recipe "配方_5": 总捻度 <- "ST_HMI_Var_HMI_r64NianDu_all", 支数 <- "ST_HMI_Var_HMI_r64ZhiShu_ChengSha", 牵伸捻度匹配值 <- "ST_HMI_Var_HMI_r64NianDu_QianShen_Best", 出车速度 <- "ST_HMI_Var_HMI_r64Velocity_ChuChe", 追捻开始捻度 <- "ST_HMI_Var_HMI_r64NianDu_1", 追捻锭子速度 <- "ST_HMI_Var_HMI_r64NianSu_2", 捻缩开始捻度 <- "ST_HMI_Var_HMI_r64NianDu_NianSuo", 捻缩距离 <- "ST_HMI_Var_HMI_r64Position_NianSuo", 追捻启用开关 <- "ST_HMI_Var_HMI_boNianDu_3"

screen "保养提示" 1280x733, template "模板_2"
   on GenerateScreen: SetTag("变量_100", 6)
   Button "HmiScreenItemData_1" at 1116,65 size 159x60; TextOn '向后 / 後向き / 뒤로'; TextOff '向后 / 後向き / 뒤로'
      on Release: ActivateScreen("自动画面", 0)
   TextField "文本域_6" at 16,8 size 995x720; Text '1.锭子油更换:每隔 天,更换一次 2.龙带传动部分12个黄油嘴，加黄油（耐高温、高速、高负荷） 3.龙带压紧器，加黄油（耐高温 、高速、高负荷） 4.弓轴滚针轴承，每年加一次黄油 5.TC龙带，每两年清洗一次，水温小于15℃，阴凉通风处晾干 6.锭子传动同步带8M-2272 检查维护 7.控制柜清洁，三个月一次,用吸吹风机来吸内部粉尘 8.锭子电机风扇绕毛清理，两个月清理一次 9.其他，走车同步带轮、走车走轮绕毛定期检查清理 1．スピンドル油交換 日,更换一次 2. タンジェントベルト伝動部12ヶ所グリスニップルに、グリス注油（耐高温・高速・高負荷） 3．タンジェントベルトのテークアップ装置にグリス注油（耐高温・高速・高負荷） 4．フォーラーシャフトのニードルベアリングに、年一回グリス注油 5．タンジェンシャルベルトを2年ごとに一回ぬるま湯（水温15℃）で洗い、かげ干しを行う。 6．スピンドル駆動タイミングベルト（８Ｍ－２２７２）点検勧奨 7．コントロールボックスを清潔にし、換気扇の粉塵を三か月ごとに吹き飛ばす。 8．锭子电机风扇绕毛清理，两个月清理一次 9．其他，走车同步带轮、走车走轮绕毛定期检查清理 1. 스핀들오일 교체: 일 간격으로 한번씩 교체한다. 2. tangential belt 전동부분12개 그리스 니플에 그리스 주입(내고온,고속,고부하) 3. 콘택트롤러에그리스 주입한다.(내고온,고속,고부하) 4. 호랑축 니들 베어링은 1년에한번씩 그리스 주입한다. 5. TCtangential belt는2년에 한번씩 청소하고 수온은 15℃이하여야 하며 서늘하고 통 풍이 잘되는곳에 말린다. 6. 스핀들 전동 타이밍벨트8M-2272를점검,유지보수한다. 7. 제어함 청소는 3개월에 한번씩 하고 흡입 송풍기로 내부 분진을 흡입한다. 8. 스핀들 모터팬감긴 원료（绕毛）청소는 2개월에 한번씩한다. 9. 기타 캐리지타이밍풀리,캐리지유동륜은정기적으로 감긴 원료(绕毛)점검,정리한다.'
   IOField "IO 域_3" at 906,98 size 65x39; FormatPattern 999
      ProcessValue <- "ST_Maintenance_g_u16_1_Times_OilChange_DingZi"
   IOField "IO 域_4" at 906,143 size 65x39; FormatPattern 999
      ProcessValue <- "ST_Maintenance_g_u16_2_Times_LongDai_HuangYouZui"
   IOField "IO 域_5" at 906,189 size 65x40; FormatPattern 999
      ProcessValue <- "ST_Maintenance_g_u16_3_Times_LongDai_YaJinQi"
   IOField "IO 域_6" at 906,236 size 65x39; FormatPattern 999
      ProcessValue <- "ST_Maintenance_g_u16_4_Times_GongZhou_Bearing"
   IOField "IO 域_7" at 906,282 size 65x39; FormatPattern 999
      ProcessValue <- "ST_Maintenance_g_u16_5_Times_LongDai_Clean"
   IOField "IO 域_8" at 906,328 size 65x40; FormatPattern 999
      ProcessValue <- "ST_Maintenance_g_u16_6_Times_DingZi_ChuanDong"
   IOField "IO 域_9" at 906,375 size 65x39; FormatPattern 999
      ProcessValue <- "ST_Maintenance_g_u16_7_Times_ControlBox_Clean"
   IOField "IO 域_10" at 906,421 size 65x39; FormatPattern 999
      ProcessValue <- "ST_Maintenance_g_u16_8_Times_DingZi_Fan"
   IOField "IO 域_1" at 258,96 size 66x39; Authorization "User administration"; FormatPattern 999
      ProcessValue <- "ST_Maintenance_g_u16_TimeInterval_OilChange"
   IOField "IO 域_2" at 486,15 size 65x39; Authorization "User administration"; FormatPattern 999
      ProcessValue <- "ST_Maintenance_g_u16_TimeReminder_Maintennance"
   TextField "文本域_4" at 334,19 size 149x32; Text '保养提醒持续 / 保全提醒 / 유지보수 알림'
   TextField "文本域_5" at 563,19 size 48x32; Text '天 / 日 / 일'
   Button "OBJECT_124" at 396,610 size 160x66; TextOn '罗拉关 / 롤러 off'; TextOff '罗拉开关 / EXIT / ローラースイッチ / 롤러 스위치'; Authorization "Operate_5"
      on Release: InvertBit("ST_Main_Var_ST_LuoLaSwitch")
      Appearance <- "ST_Main_Var_ST_LuoLaSwitch"
   TextField "文本域_1" at 40,56 size 149x32; Text '保养项目 / 保全項目 / 유지보수 항목'
   TextField "文本域_2" at 850,56 size 149x32; Text '保养次数 / 保全回数 / 유지보수 횟수'

screen "报警画面" 1280x733, template "模板_2"
   on GenerateScreen: SetTag("变量_100", 5)
   Button "HmiScreenItemData_1" at 1112,90 size 159x60; TextOn '向后 / 後向き / 뒤로'; TextOff '向后 / 後向き / 뒤로'
      on Release: function_efd93a16()
   Button "HmiScreenItemData_2" at 1112,224 size 159x60; TextOn '向后 / 後向き / 뒤로'; TextOff '报警记录 / 警報記録 / 경보알람기록'
      on Release: ActivateScreen("报警记录", 0)
   Button "HmiScreenItemData_3" at 1112,360 size 159x60; TextOn '向后 / 後向き / 뒤로'; TextOff '自动画面 / 自動画面 / 자동화면'
      on Release: ActivateScreen("自动画面", 0)
   AlarmView "报警视图_1" at 3,3 size 1101x728

screen "报警记录" 1280x733, template "模板_2"
   on GenerateScreen: SetTag("变量_100", 16)
   AlarmView "报警视图_1" at 3,2 size 1105x729; ColumnTextDevice 'D425 / PLC / API / ПЛК'
   Button "HmiScreenItemData_2" at 1118,71 size 159x60; TextOn '向后 / 後向き / 뒤로'; TextOff '向后 / 後向き / 뒤로'
      on Release: ActivateScreen("报警画面", 0)

screen "生头画面" 1280x733, template "模板_2"
   on GenerateScreen: SetTag("变量_100", 4)
   Button "HmiScreenItemData_1" at 1118,192 size 159x60; TextOn '向后 / 後向き / 뒤로'; TextOff '向后 / 後向き / 뒤로'
      on Release: ActivateScreen("自动画面", 0)
   Button "OBJECT_107" at 864,104 size 200x65; TextOff '手动 / EXIT / 手動 / 수동'
      on Press: SetTag("ST_Main_Var_g_i16_Mode_Selected", 4)
      Appearance <- "ST_Main_Var_g_bo_Mode_Enabled_Manual"
   Button "OBJECT_108" at 864,192 size 200x65; TextOff '空锭(先插管) EXIT 空鍾（糸管挿入済み） 아이들 스핀들 (먼저 보빈관을 삼입)'
      on Release: ResetBit("ST_HMI_Var_HMI_bo_KongDingShengTou")
      on Press: SetBit("ST_HMI_Var_HMI_bo_KongDingShengTou")
      Appearance <- "ST_HMI_Var_HMI_i16_ShengTou_Select"
   Button "OBJECT_106" at 1041,4 size 238x39; TextOff '手动 / EXIT / 手動 / 수동'; TextList "mode_enabled_1"
      ProcessValue <- "ST_Main_Var_g_i16_Mode_Enabled"
      Appearance <- "ST_Main_Var_g_i16_Mode_Enabled"
   TextField "Text Field_45" at 370,139 size 151x47; Text '实际牵伸: / 実際ドラフト: / 실제 드라프트:'
   TextField "Text Field_46" at 370,205 size 151x47; Text '分散牵伸: / 分散ドラフト: / 스핀들 드라프트:'
   TextField "Text Field_47" at 370,270 size 151x47; Text '走车位置: / キャレージ位置: / 캐리지위치:'
   Button "OBJECT_111" at 1041,43 size 238x40; TextOff '手动 / EXIT / 手動 / 수동'; TextList "KongDing_status#mig1"
      Visibility <- "ST_Main_Var_g_bo_Mode_Enabled_KongDing"
      ProcessValue <- "ST_Main_Var_g_i16_KongDing_Status"
      Appearance <- "ST_Main_Var_g_i16_KongDing_Status"
   Button "OBJECT_109" at 864,456 size 200x66; TextOff '启动 / EXIT / 起動 / 가동'
      on Release: ResetBit("ST_HMI_Var_HMI_bo_ShengTou_QiDong")
      on Press: SetBit("ST_HMI_Var_HMI_bo_ShengTou_QiDong")
      Visibility <- "ST_Main_Var_g_i16_Mode_Enabled"
      Appearance <- "ST_Main_Var_g_bo_KongDing_Running_Status"
   Button "OBJECT_110" at 864,544 size 200x65; TextOff '停止 / EXIT / 정지'
      on Release: ResetBit("ST_HMI_Var_HMI_bo_ShengTou_TingZhi")
      on Press: SetBit("ST_HMI_Var_HMI_bo_ShengTou_TingZhi")
      Visibility <- "ST_Main_Var_g_i16_Mode_Enabled"
      Appearance <- "ST_Main_Var_g_bo_KongDing_Running_Status"
   TextField "Text Field_49" at 167,635 size 125x39; Text '单纱张力 / 単糸張力 / 단사 장력'
   TextField "Text Field_50" at 40,635 size 127x39; Text '纱穗个数 / コップ本数: / 코프갯수'
   TextField "Text Field_51" at 292,635 size 252x39; Text '总张力目标值|实时值 / 総張力目標値|実際値 / 전체 장력 목표값| 실시간값'
   TextField "Text Field_52" at 544,635 size 253x39; Text '弓位置目标值|实时值 / フォーラー位置目標値|実際値 / 호랑위치 목표값 |실시간값'
   TextField "Text Field_72" at 40,596 size 757x39; Text '张力控制 / 巻取張力制御 / 장력 제어'
   TextField "Text Field_53" at 370,74 size 151x47; Text '实际捻度: / 実際撚数： / 실제연도:'
   Button "OBJECT_112" at 864,368 size 200x66; TextOff '落纱生头 / EXIT / 玉揚げ口付け / 돕핑스레드업'
      on Release: ResetBit("ST_HMI_Var_HMI_bo_LuoShaShengTou")
      on Press: SetBit("ST_HMI_Var_HMI_bo_LuoShaShengTou")
      Appearance <- "ST_HMI_Var_HMI_i16_ShengTou_Select"
   TextField "Text Field_54" at 643,90 size 16x27; Text '/'
   TextField "Text Field_55" at 643,155 size 16x27; Text '/'
   TextField "Text Field_56" at 643,221 size 16x27; Text '/'
   TextField "Text Field_2" at 40,74 size 169x45; Text '总捻度: / 総撚数： / 전체 연도:'
   TextField "Text Field_25" at 40,139 size 169x45; Text '总牵伸: / 総ドラフト: / 전체 드라프트:'
   TextField "Text Field_26" at 40,270 size 169x46; Text '送条牵伸: / 篠送出しドラフト: / 시누 공급드라프트:'
   TextField "Text Field_27" at 40,205 size 169x45; Text '分散牵伸: / 分散ドラフト: / 스핀들 드라프트:'
   TextField "Text Field_57" at 370,466 size 151x47; Text '成形位置: / コップ形成位置: / 성형 위치:'
   TextField "Text Field_58" at 370,531 size 151x47; Text '张力位置: / 張力位置: / 장력 위치:'
   TextField "Text Field_59" at 370,336 size 151x47; Text '罗拉位置: / ローラー位置: / 롤러 위치:'
   TextField "Text Field_60" at 370,400 size 151x47; Text '滚筒位置: / ターンポール位置: / 시누공급 길이:'
   TextField "Text Field_14" at 86,21 size 196x39; Text '设定参数显示 / 設定パラメーター表示 / 매개변수 설정'
   IOField "IO Field_28" at 531,139 size 112x45; FormatPattern 9.99
      ProcessValue <- "ST_HMI_Var_HMI_r64QianShen_All_real_ShengTou"
   IOField "IO Field_29" at 531,205 size 112x45; FormatPattern 99.99
      ProcessValue <- "ST_HMI_Var_HMI_r64QianShen_FenSan_real_ShengTou"
   IOField "IO Field_30" at 531,270 size 112x46; FormatPattern 9999
      ProcessValue <- "ST_HMI_Var_HMI_r64Axis_ZouChe_Position_real"
   TextField "Text Field_15" at 502,21 size 196x39; Text '实时参数显示 / 実際パラメーター表示: / 실시간 매개변수 표시'
   IOField "IO Field_75" at 40,674 size 127x40; FormatPattern 9999
      ProcessValue <- "ST_HMI_Var_HMI_r64_ShuLiang_ShaSui"
   IOField "IO Field_76" at 167,674 size 125x40; FormatPattern 999.9
      ProcessValue <- "ST_HMI_Var_HMI_r64_DanSha_ZhangLi_ShengTou"
   IOField "IO Field_77" at 292,674 size 127x40; FormatPattern 999.99
      ProcessValue <- "ST_Main_Var_g_r64Axis_1_ZhangLi_Torque_Limit_Positive"
   IOField "IO Field_78" at 419,674 size 125x40; FormatPattern 999.99
      ProcessValue <- "Axis_1_ZhangLi_torqueLimitPositive_value"
   IOField "IO Field_79" at 544,674 size 127x40; FormatPattern 999.9
      ProcessValue <- "ST_HMI_Var_HMI_r64Axis_1_ZhangLi_Position_JuanRao_Set_KongDing_12"
   IOField "IO Field_80" at 671,674 size 126x40; FormatPattern 999.9
      ProcessValue <- "ST_HMI_Var_HMI_r64Axis_1_ZhangLi_Position_JuanRao_real"
   IOField "IO Field_32" at 531,74 size 112x45; FormatPattern 9999
      ProcessValue <- "ST_HMI_Var_HMI_r64NianDu_real_ShengTou"
   IOField "IO Field_43" at 671,74 size 112x45; FormatPattern 9999
      on OnFinishInput: SetBit("ST_Calculation_Var_HMI_bo_Calculation_0_Start"); SetTag("ST_Calculation_Var_g_i16_Calculation_0_3_Select_Status", 1)
      ProcessValue <- "ST_HMI_Var_HMI_r64NianDu_all"
   IOField "IO Field_14" at 671,139 size 112x45; FormatPattern 9.99
      ProcessValue <- "ST_HMI_Var_HMI_r64QianShen_All_KongDing_7"
   IOField "IO Field_16" at 671,205 size 112x45; FormatPattern 9.99
      ProcessValue <- "ST_HMI_Var_HMI_r64QianShen_FenSan_KongDing_7"
   IOField "IO Field_44" at 221,74 size 112x45; FormatPattern 9999
      on OnFinishInput: SetBit("ST_Calculation_Var_HMI_bo_Calculation_0_Start"); SetTag("ST_Calculation_Var_g_i16_Calculation_0_3_Select_Status", 1)
      ProcessValue <- "ST_HMI_Var_HMI_r64NianDu_all"
   IOField "IO Field_15" at 219,139 size 112x45; FormatPattern 9.99
      ProcessValue <- "ST_HMI_Var_HMI_r64QianShen_All"
   IOField "IO Field_17" at 219,270 size 112x46; FormatPattern 9.999
      ProcessValue <- "ST_HMI_Var_HMI_r64QianShen_WuNian"
   IOField "IO Field_18" at 219,205 size 112x45; FormatPattern 9.99
      ProcessValue <- "ST_HMI_Var_HMI_r64QianShen_FenSan"
   IOField "IO Field_74" at 531,466 size 112x46; FormatPattern 99.9
      ProcessValue <- "ST_HMI_Var_HMI_r64Axis_ChengXing_Position_real"
   IOField "IO Field_82" at 531,531 size 112x47; FormatPattern 99.9
      ProcessValue <- "ST_HMI_Var_HMI_r64Axis_1_ZhangLi_Position_JuanRao_real"
   IOField "IO Field_33" at 531,400 size 112x47; FormatPattern 9999
      ProcessValue <- "Axis_GunTong_positioningState_actualPosition"
   IOField "IO Field_66" at 531,336 size 112x45; FormatPattern 9999
      ProcessValue <- "Axis_LuoLa_positioningState_actualPosition"
   TextField "Text Field_29" at 40,336 size 169x45; Text '速度比例: / 속도비율:'
   TextField "Text Field_62" at 40,398 size 169x45; Text '出车展距: / 出機展開距離: / 외진거리:'
   IOField "IO Field_19" at 219,336 size 112x45; FormatPattern 9.99
      ProcessValue <- "ST_HMI_Var_HMI_r64_Scale_KongDing_7"
   IOField "IO Field_35" at 219,400 size 112x47; FormatPattern 9999
      ProcessValue <- "ST_HMI_Var_HMI_r64Position_ChuChe_KongDing_7"
   Button "OBJECT_3" at 824,643 size 160x71; TextOff '标准纱管1 / EXIT / 標準糸管１ / 표준보빈1'; Authorization "Monitor"
      on Press: SetTag("ST_HMI_Var_HMI_i16_Status_ShaGuan_Select", 1)
      Appearance <- "ST_HMI_Var_HMI_i16_Status_ShaGuan_Select"
   Button "OBJECT_4" at 1008,643 size 160x71; TextOff '标准纱管2 / EXIT / 標準糸管２ / 표준보빈2'; Authorization "Monitor"
      on Press: SetTag("ST_HMI_Var_HMI_i16_Status_ShaGuan_Select", 2)
      Appearance <- "ST_HMI_Var_HMI_i16_Status_ShaGuan_Select"
   Button "OBJECT_5" at 864,280 size 200x65; TextOff '空锭(光锭) EXIT 空鍾 아이들 스핀들 (광스핀들)'
      on Release: ResetBit("ST_HMI_Var_HMI_bo_KongDingShengTou_GuangDing")
      on Press: SetBit("ST_HMI_Var_HMI_bo_KongDingShengTou_GuangDing")
      Appearance <- "ST_HMI_Var_HMI_i16_ShengTou_Select"
   Button "OBJECT_1" at 1104,367 size 173x66; TextOff '拔锭脚纱选择 / EXIT / 시다구미'
      on Release: InvertBit("ST_HMI_Var_HMI_bo_BaShaTou_Select")
      Appearance <- "ST_HMI_Var_HMI_bo_BaShaTou_Select"
      Visibility <- "ST_HMI_Var_HMI_i16_ShengTou_Select"
      ObjectEnable <- "ST_Main_Var_g_i16_KongDing_Status"
   IOField "IO Field_1" at 219,466 size 112x47; FormatPattern 99
      ProcessValue <- "ST_HMI_Var_HMI_r64Axis_ZouChe_Position_LuoSha_112_Delta_BaTou"
   TextField "Text Field_1" at 40,467 size 169x46; Text '拔锭脚纱补偿距离: / 拔锭脚纱补偿距离:: / 시다구미 거리'

screen "时间显示" 1280x733, template "模板_2"
   on GenerateScreen: SetTag("变量_100", 7); "timeConverse"()
   Button "按钮_1" at 174,88 size 95x82; TextOn '出车 / 出機 / 외진'; TextOff '出车 / 出機 / 외진'
      Appearance <- "ST_Main_Var_g_i16_Automatic_Status"
   Button "按钮_2" at 321,88 size 95x82; TextOn '加捻 / 撚掛 / 연사'; TextOff '加捻 / 撚掛 / 연사'
      Appearance <- "ST_Main_Var_g_i16_Automatic_Status"
   Button "按钮_3" at 457,88 size 117x82; TextOn '退绕 パッキン グオフ 언와인딩'; TextOff '退绕 パッキン グオフ 언와인딩'
      Appearance <- "ST_Main_Var_g_i16_Automatic_Status"
   Button "按钮_4" at 614,88 size 95x82; TextOn '进车 / 入機 / 내진'; TextOff '进车 / 入機 / 내진'
      Appearance <- "ST_Main_Var_g_i16_Automatic_Status"
   Button "按钮_5" at 760,88 size 96x82; TextOn '周期 / サイクル / 주기'; TextOff '周期 / サイクル / 주기'
      Appearance <- "ST_Main_Var_g_i16_Automatic_Status"
   TextField "文本域_1" at 33,356 size 274x31; Text '系统总运行时间: / システム総運転時間: / 시스템 전체 운행 시간'
   TextField "文本域_2" at 400,356 size 31x31; Text '年 / 년'
   TextField "文本域_4" at 514,356 size 31x31; Text '天 / 日 / 일'
   TextField "文本域_5" at 617,356 size 31x31; Text '时 / 時 / 시'
   TextField "文本域_6" at 715,356 size 31x31; Text '分 / 분'
   TextField "文本域_7" at 814,356 size 31x31; Text '秒 / 초'
   IOField "IO Field_23" at 174,183 size 95x55; FormatPattern 99.99
      ProcessValue <- "ST_Main_Var_g_r64_Time_chuche"
   IOField "IO Field_24" at 321,183 size 95x55; FormatPattern 99.99
      ProcessValue <- "ST_Main_Var_g_r64_Time_jianian"
   IOField "IO Field_25" at 467,183 size 96x55; FormatPattern 99.99
      ProcessValue <- "ST_Main_Var_g_r64_Time_tuirao"
   IOField "IO Field_26" at 614,183 size 95x55; FormatPattern 99.99
      ProcessValue <- "ST_Main_Var_g_r64_Time_juanrao"
   IOField "IO Field_27" at 760,183 size 96x55; FormatPattern 99.99
      ProcessValue <- "ST_Main_Var_g_r64_Time_Once"
   IOField "IO Field_29" at 323,346 size 72x55; FormatPattern 999
      ProcessValue <- "VBS_time_year"
   IOField "IO Field_30" at 439,346 size 68x55; FormatPattern 999
      ProcessValue <- "VBS_time_day"
   IOField "IO Field_30#mig1" at 553,346 size 55x55; FormatPattern 99
      ProcessValue <- "VBS_time_hour"
   IOField "IO Field_31" at 654,346 size 55x55; FormatPattern 99
      ProcessValue <- "VBS_time_min"
   IOField "IO Field_32" at 755,346 size 52x55; FormatPattern 99
      ProcessValue <- "VBS_time_sec"
   Button "HmiScreenItemData_1" at 1116,65 size 159x60; TextOn '向后 / 後向き / 뒤로'; TextOff '向后 / 後向き / 뒤로'
      on Release: ActivateScreen("自动画面", 0)

screen "自动画面" 1280x733
   on GenerateScreen: SetTag("变量_100", 1)
   Button "HmiScreenItemData_7" at 1118,670 size 159x57; TextOff 'Text'; Authorization "Operate_4"
      on Release: ActivateScreen("常用调试画面", 0); ResetBit("HMI_Tag_bo_showDebugButton")
      ObjectEnable <- "HMI_Tag_bo_showDebugButton"
   Button "HmiScreenItemData_1" at 1118,112 size 159x60; TextOn '手动画面 / 手動画面 / 수동화면'; TextOff '手动画面 / 手動画面 / 수동화면'
      on Release: ActivateScreen("手动画面", 0)
   Button "HmiScreenItemData_2" at 1118,395 size 159x60; TextOn '报警画面 / Alarm Pic / 警報画面 / 경보화면'; TextOff '报警画面 / Alarm Pic / 警報画面 / 경보화면'
      on Release: ActivateScreen("报警画面", 0)
   Button "HmiScreenItemData_4" at 1118,206 size 159x60; TextOn '设置画面 / 設置画面 / 설정화면'; TextOff '设置画面 / 設置画面 / 설정화면'
      on Release: ActivateScreen("设置画面", 0); ResetBit("HMI_Tag_bo_showDebugButton")
   Button "HmiScreenItemData_5" at 1118,490 size 159x60; TextOn '保养提示 / MAINTENANCE ALERT / 保全画面 / 유지보수 알림'; TextOff '保养提示 / MAINTENANCE ALERT / 保全画面 / 유지보수 알림'
      on Release: ActivateScreen("保养提示", 0)
   Button "HmiScreenItemData_6" at 1118,585 size 159x60; TextOn '时间显示 / 時間表示 / 시간표시'; TextOff '时间显示 / 時間表示 / 시간표시'
      on Release: ActivateScreen("时间显示", 0)
   Button "HmiScreenItemData_9" at 1118,301 size 159x60; TextOn '生头画面 / 生頭画面 / 스레드업화면'; TextOff '生头画面 / 生頭画面 / 스레드업화면'
      on Release: ActivateScreen("生头画面", 0)
   TextField "Text Field_19" at 0,64 size 126x42; Text '纺纱批数 / 紡績ロット数 / 방적 로트'
   TextField "Text Field_22" at 126,64 size 126x42; Text '累计亨司 / 累計 Hanks / 누계횟수'
   TextField "Text Field_23" at 253,65 size 126x42; Text '本次亨司 / 今回 Hanks / 당차횟수'
   TextField "Text Field_28" at 0,148 size 126x42; Text '实时跟踪 / リアルタイム 追跡 / 실시간 추적'
   TextField "Text Field_29" at 126,148 size 126x42; Text '走车位置 / CarriagePos / キャレージ位置 / 캐리지위치'
   TextField "Text Field_30" at 252,148 size 126x42; Text '捻度 / 撚数 / 연도'
   TextField "Text Field_31" at 378,148 size 126x42; Text '锭子速度 / スピンドル回転数 / 스핀들속도'
   TextField "Text Field_32" at 504,148 size 126x42; Text '总牵伸 / draft / 総ドラフト / 전체 드라프트'
   TextField "Text Field_33" at 630,148 size 126x42; Text '分散牵伸 / 分散ドラフト / 스핀들 드라프트'
   TextField "Text Field_34" at 756,148 size 126x42; Text '送条长度 / 篠送り出し長 / 시누공급길이'
   TextField "Text Field_35" at 0,190 size 126x42; Text '目标值 / 目標値 / 목표값'
   TextField "Text Field_36" at 0,232 size 126x42; Text '设定值 / 実際値 / 설정값'
   TextField "Text Field_38" at 0,22 size 882x42; Text '系统运行情况 / System Running State / システム運転状況 / 시스템 운행 상황'
   TextField "Text Field_39" at 252,334 size 126x42; Text '起始点高度 / 開始点高度 / 출발점 높이'
   TextField "Text Field_40" at 126,334 size 126x42; Text '成纱支数 / 番手: / 실 번수'
   TextField "Text Field_41" at 378,334 size 126x42; Text '下锥体高度 / 下錐体高度 / 하단코프높이'
   TextField "Text Field_42" at 504,334 size 126x42; Text '上锥体高度 / 上錐体高度 / 상단 코프높이'
   TextField "Text Field_43" at 630,334 size 126x42; Text '最大直径 / MaxDiameter / 최대 직경'
   TextField "Text Field_44" at 756,334 size 126x42; Text '实时位置 / 実際位置 / 실시간값'
   TextField "Text Field_45" at 0,334 size 126x42; Text '纱穗参数 / コップ数 / 코프 형성'
   TextField "Text Field_46" at 0,376 size 126x42; Text '设定值 / 設定値 / 설정값'
   Button "OBJECT_106" at 884,0 size 238x42; TextOff '手动 / EXIT / 手動 / 수동'; TextList "mode_enabled_1"
      ProcessValue <- "ST_Main_Var_g_i16_Mode_Enabled"
      Appearance <- "ST_Main_Var_g_i16_Mode_Enabled"
   Button "OBJECT_107" at 910,112 size 182x70; TextOff '手动 / EXIT / 手動 / 수동'
      on Press: SetTag("ST_Main_Var_g_i16_Mode_Selected", 4)
      Appearance <- "ST_Main_Var_g_i16_Manual_Status"
   Button "OBJECT_108" at 910,217 size 182x70; TextOff '自动 / Auto / 自動 / 자동'
      on Release: ResetBit("ST_HMI_Var_HMI_bo_Auto")
      on Press: SetBit("ST_HMI_Var_HMI_bo_Auto")
      Appearance <- "ST_Main_Var_g_bo_Mode_Enabled_Automatic"
   Button "OBJECT_109" at 910,323 size 182x70; TextOff '启动 / EXIT / 起動 / 가동'
      on Press: SetBit("ST_Main_Var_g_bo_Automatic_Running_Selected")
      Visibility <- "ST_Main_Var_g_bo_Mode_Enabled_Automatic"
      Appearance <- "ST_Main_Var_g_bo_Automatic_Running_Status"
   Button "OBJECT_110" at 910,428 size 182x70; TextOff '停止 / 정지'
      on Press: SetTag("ST_Main_Var_g_i16_Automatic_Stopping_Selected", 1)
      Visibility <- "ST_Main_Var_g_bo_Mode_Enabled_Automatic"
      Appearance <- "ST_Main_Var_g_i16_Automatic_Stopping_Selected"
   TextField "Text Field_47" at 252,476 size 126x42; Text '单纱张力 / 単糸張力 / 단사 장력'
   TextField "Text Field_48" at 126,476 size 126x42; Text '纱穗个数 / コップ本数 / 코프갯수'
   TextField "Text Field_49" at 378,476 size 252x42; Text '总张力目标值|实时值 / 総張力目標値|実際値 / 전체 장력 목표값| 실시간값'
   TextField "Text Field_50" at 630,476 size 252x42; Text '弓位置目标值|实时值 / フォーラー位置目標値|実際値 / 호랑위치 목표값 |실시간값'
   TextField "Text Field_53" at 0,476 size 126x42; Text '纱穗参数 / コップ数 / 코프 매개변수'
   TextField "Text Field_54" at 0,518 size 126x42; Text '设定值 / 設定値 / 설정값'
   TextField "Text Field_71" at 1,292 size 881x42; Text '成形控制 / コップ形成制御 / 성형제어'
   TextField "Text Field_72" at 0,434 size 882x42; Text '张力控制 / 巻取張力制御 / 장력 제어'
   Button "OBJECT_111" at 884,43 size 238x42; TextOff '手动 / EXIT / 手動 / 수동'; TextList "automatic_status_1"
      Visibility <- "ST_Main_Var_g_bo_Mode_Enabled_Automatic"
      ProcessValue <- "ST_Main_Var_g_i16_Automatic_Status"
      Appearance <- "ST_Main_Var_g_i16_Automatic_Status"
   Button "OBJECT_112" at 250,654 size 126x56; TextOff '出车 / EXIT / 出機 / 외진'; Authorization "User administration"
      on Press: SetTag("ST_Main_Var_g_i16_Automatic_Selected", 8); function_f23ef4c9()
      Appearance <- "ST_Main_Var_g_i16_Automatic_Selected"
   Button "OBJECT_113" at 376,654 size 126x56; TextOff '出车到 / EXIT / 出機完了 / 외진도착'; Authorization "User administration"
      on Press: SetTag("ST_Main_Var_g_i16_Automatic_Selected", 16); function_f23ef4c9()
      Appearance <- "ST_Main_Var_g_i16_Automatic_Selected"
   Button "OBJECT_114" at 502,654 size 126x56; TextOff '退绕 / パッキングオフ / 언와인딩'; Authorization "User administration"
      on Press: SetTag("ST_Main_Var_g_i16_Automatic_Selected", 32); function_f23ef4c9()
      Appearance <- "ST_Main_Var_g_i16_Automatic_Selected"
   Button "OBJECT_115" at 628,654 size 126x56; TextOff '卷绕 / EXIT / 巻取 / 와인딩'; Authorization "User administration"
      on Press: SetTag("ST_Main_Var_g_i16_Automatic_Selected", 64); function_f23ef4c9()
      Appearance <- "ST_Main_Var_g_i16_Automatic_Selected"
   Button "OBJECT_116" at 754,654 size 126x56; TextOn '存绕 / 逆巻取 / 와인딩 저장'; TextOff '存绕 / EXIT / 逆巻取 / 와인딩 저장'; Authorization "User administration"
      on Press: SetTag("ST_Main_Var_g_i16_Automatic_Selected", 128); function_f23ef4c9()
      Appearance <- "ST_Main_Var_g_i16_Automatic_Selected"
   Button "OBJECT_117" at 910,534 size 182x70; TextOff '紧急停止 / EXIT / 緊急停止 / 비상정지'
      on Press: SetTag("ST_Main_Var_g_i16_Automatic_Selected", 2)
   Button "OBJECT_118" at 910,640 size 182x70; TextOff '退出紧急停止 / 緊急停止を終了する / 비상정지종료'
      on Press: SetTag("ST_Main_Var_g_i16_Automatic_Status", 1)
      Visibility <- "ST_Main_Var_g_bo_Automatic_Status_Mergestop"
   TextField "文本域_1" at 154,581 size 70x42; Text 'sec'
   TextField "文本域_2" at 154,639 size 94x42; Text 'm/min'
   IOField "IO Field_44" at 126,106 size 126x42; FormatPattern 99999999
      ProcessValue <- "ST_Main_Var_g_u32_N_Cycle_Whole"
   IOField "IO Field_45" at 252,106 size 126x42; FormatPattern 9999
      ProcessValue <- "ST_Main_Var_g_u16_N_Cycle_Single"
   IOField "IO Field_50" at 126,190 size 126x42; FormatPattern 9999.9
      ProcessValue <- "ST_HMI_Var_HMI_r64Axis_ZouChe_Position_object"
   IOField "IO Field_51" at 126,232 size 126x42; FormatPattern 9999.9
      ProcessValue <- "ST_HMI_Var_HMI_r64Axis_ZouChe_Position_real"
   IOField "IO Field_53" at 252,190 size 126x42; FormatPattern 9999
      ProcessValue <- "ST_HMI_Var_HMI_r64Niandu_all_Current"
   IOField "IO Field_54" at 252,232 size 126x42; FormatPattern 9999
      ProcessValue <- "ST_HMI_Var_HMI_r64NianDu_real"
   IOField "IO Field_56" at 378,190 size 126x42; FormatPattern 99999
      ProcessValue <- "ST_HMI_Var_HMI_r64Axis_DingZi_Velocity_object"
   IOField "IO Field_57" at 378,232 size 126x42; FormatPattern 99999
      ProcessValue <- "ST_HMI_Var_HMI_r64Axis_DingZi_Velocity_real"
   IOField "IO Field_59" at 504,190 size 126x42; FormatPattern 9.99
      ProcessValue <- "ST_HMI_Var_HMI_r64QianShen_All"
   IOField "IO Field_60" at 504,232 size 126x42; FormatPattern 9.999
      ProcessValue <- "ST_HMI_Var_HMI_r64QianShen_All_real"
   IOField "IO Field_62" at 630,190 size 126x42; FormatPattern 9.99
      ProcessValue <- "ST_HMI_Var_HMI_r64QianShen_FenSan"
   IOField "IO Field_63" at 630,232 size 126x42; FormatPattern 99.999
      ProcessValue <- "ST_HMI_Var_HMI_r64QianShen_FenSan_real"
   IOField "IO Field_65" at 756,190 size 126x42; FormatPattern 9999.9
      ProcessValue <- "ST_Main_Var_g_r64Axis_LuoLa_Position"
   IOField "IO Field_66" at 756,232 size 126x42; FormatPattern 9999.9
      ProcessValue <- "Axis_LuoLa_positioningState_commandPosition"
   IOField "IO Field_68" at 1,106 size 126x42; FormatPattern 9999
      ProcessValue <- "ST_Main_Var_g_u16_PiShu_Whole"
   IOField "IO Field_69" at 126,376 size 126x42; FormatPattern 99.99
      ProcessValue <- "ST_HMI_Var_HMI_r64ZhiShu_ChengSha"
   IOField "IO Field_70" at 252,376 size 126x42; FormatPattern 99.9
      ProcessValue <- "ST_HMI_Var_HMI_r64Height_ShaSui_Start"
   IOField "IO Field_71" at 378,376 size 126x42; FormatPattern 99.9
      ProcessValue <- "ST_HMI_Var_HMI_r64Height_ShaSui_Bottom"
   IOField "IO Field_72" at 504,376 size 126x42; FormatPattern 99.9
      ProcessValue <- "ST_HMI_Var_HMI_r64Height_ShaSui_Top"
   IOField "IO Field_74" at 756,376 size 126x42; FormatPattern 99.9
      ProcessValue <- "ST_HMI_Var_HMI_r64Axis_ChengXing_Position_real"
   IOField "IO Field_77" at 378,518 size 126x42; FormatPattern 999.99
      ProcessValue <- "ST_Main_Var_g_r64Axis_1_ZhangLi_Torque_Limit_Positive"
   IOField "IO Field_78" at 504,518 size 126x42; FormatPattern 999.99
      ProcessValue <- "Axis_1_ZhangLi_torqueLimitPositive_value"
   IOField "IO Field_79" at 630,518 size 126x42; FormatPattern 999.9
      ProcessValue <- "ST_VAR_ZhangLi_g_r64Axis_1_ZhangLi_Position_JuanRao_Set"
   IOField "IO Field_80" at 756,518 size 126x42; FormatPattern 999.9
      ProcessValue <- "ST_HMI_Var_HMI_r64Axis_1_ZhangLi_Position_JuanRao_real"
   IOField "IO Field_81" at 18,581 size 126x42; FormatPattern 999.9999
      ProcessValue <- "ST_Main_Var_g_r64_Time_Once"
   IOField "IO Field_82" at 18,640 size 126x42; FormatPattern 999.9999
      ProcessValue <- "ST_Main_Var_g_r64_Length_One_Minute"
   IOField "IO Field_83" at 630,376 size 126x42; FormatPattern 99.9
      ProcessValue <- "ST_HMI_Var_HMI_r64Diameter_ShaSui_Max"
   Button "按钮_2" at 0,2 size 248x42; TextOff '保养提示已隐藏 / 유지보수 알림을 이미 숨김'
      on Click: ResetBit("VBS_alwaysFalse")
      Visibility <- "VBS_alwaysFalse"
   TextField "Text Field_1" at 379,65 size 125x41; Text '满纱周期 / CarriageVelo / キャレージ速度 / 코프완성주기'
   IOField "IO Field_1" at 378,106 size 126x42; FormatPattern 9999
      ProcessValue <- "ST_FC_Var_g_N"
   Button "HmiScreenItemData_3" at 2,667 size 143x60; TextOff 'Text'
      on Release: SetBit("HMI_Tag_bo_showDebugButton")
   TextField "Text Field_2" at 505,65 size 125x41; Text '产量kg / 篠送り出し速度 / 생산량kg'
   TextField "Text Field_24" at 631,65 size 126x42; Text '纱穗重量g / RunningMode / 運転モード / 코프중량'
   TextField "Text Field_25" at 757,65 size 126x42; Text '自动状态 / AutoStatus / 自動状態 / 자동 상태'
   Button "OBJECT_121" at 757,106 size 126x42; TextOff '手动 / EXIT / 手動 / 수동'; TextList "automatic_status_2"
      Visibility <- "ST_Main_Var_g_bo_Mode_Enabled_Automatic"
      ProcessValue <- "ST_Main_Var_g_i16_Automatic_Status"
      Appearance <- "ST_Main_Var_g_i16_Automatic_Status"
   IOField "IO Field_2" at 504,106 size 126x42; FormatPattern 9999999
      ProcessValue <- "ST_Maintenance_HMI_r64_Production_Once"
   Button "OBJECT_1" at 1118,667 size 159x66; TextOff '抬 弓 / EXIT / 호랑올림'
      on Release: InvertBit("ST_MotionTask_ZhangLi_Var_HMI_bo_TaiGong")
      Appearance <- "ST_MotionTask_ZhangLi_Var_HMI_bo_TaiGong"
      ObjectEnable <- "ST_Main_Var_g_i16_Automatic_Status"
      Visibility <- "ST_Main_Var_g_i16_Mode_Enabled"
   TextField "Text Field_62" at 375,586 size 129x45; Text '放下位置: / 캐리지위치'
      Visibility <- "ST_MotionTask_ZhangLi_Var_HMI_bo_TaiGong"
   IOField "IO Field_35" at 504,585 size 126x47; FormatPattern 9999
      Visibility <- "ST_MotionTask_ZhangLi_Var_HMI_bo_TaiGong"
      ProcessValue <- "ST_MotionTask_ZhangLi_Var_HMI_r64Axis_ZouChe_Position_TaiGong_FangXia"
   IOField "IO Field_4" at 754,585 size 126x47; FormatPattern 99
      Visibility <- "ST_MotionTask_ZhangLi_Var_HMI_bo_TaiGong"
      ProcessValue <- "ST_MotionTask_ZhangLi_Var_HMI_r64Axis_1_ZhangLi_Position_TaiGong"
   TextField "Text Field_3" at 630,586 size 126x46; Text '抬弓角度: / 拔锭脚纱补偿距离:: / 호랑각도'
      Visibility <- "ST_MotionTask_ZhangLi_Var_HMI_bo_TaiGong"
   IOField "IO Field_76" at 253,517 size 126x42; FormatPattern 999.9
      ProcessValue <- "ST_HMI_Var_HMI_r64_LuoSha_Force_DanSha_ZhangLi_FangKai"
   IOField "IO Field_75" at 126,517 size 126x42; FormatPattern 9999
      ProcessValue <- "ST_HMI_Var_HMI_r64_ShuLiang_ShaSui"
   IOField "IO Field_5" at 631,107 size 126x42; FormatPattern 9999999
      ProcessValue <- "ST_Maintenance_HMI_r64_Weight_ShaSui"
   Button "HmiScreenItemData_8" at 1118,25 size 159x60; TextOn '用户管理'; TextOff '用户管理'
      on Release: ActivateScreen("用户管理", 0)
   TextField "文本域_3" at 30,98 size 812x98; Text '保养时间到,请停机第 次更换锭子 油! 保养时间到,请停机第 次更换锭子 油! 유지보수시간. 기계 스톱. 제 차 스핀들오일 교체 !'
      Visibility <- "ST_Maintenance_g_bo_1_Warn_Status_OilChange_DingZi"
   IOField "IO Field_86" at 334,100 size 70x31; FormatPattern 999
      Visibility <- "ST_Maintenance_g_bo_1_Warn_Status_OilChange_DingZi"
      ProcessValue <- "ST_Maintenance_g_u16_1_Times_TiShi_OilChange_DingZi"
   Button "按钮_1" at 597,98 size 196x42; TextOff '1小时后提醒 / 1시간후 다시 알림'
      Visibility <- "ST_Maintenance_g_bo_1_Warn_Status_OilChange_DingZi"
      on Click: ResetBit("ST_Maintenance_g_bo_1_Warn_Status_OilChange_DingZi")
   Button "按钮_3" at 597,154 size 196x42; TextOff '已保养完毕 / 유지보수 이미 완료'; Authorization "User administration"
      Visibility <- "ST_Maintenance_g_bo_1_Warn_Status_OilChange_DingZi"
      on Click: ResetBit("ST_Maintenance_g_bo_1_Status_OilChange_DingZi")
   TextField "文本域_4" at 39,105 size 812x100; Text '保养时间到,请停机第 次为龙带传动 部分黄油嘴加注黄油 保养时间到,请停机第 次为龙带传动 部分黄油嘴加注黄油 유지보수시간. 기계 스톱. 제 차 tangential belt 전동 부분 그리스 니플에 그리스를 주입한다.'
      Visibility <- "ST_Maintenance_g_bo_2_Warn_Status_LongDai_HuangYouZui"
   IOField "IO Field_87" at 345,106 size 70x29; FormatPattern 999
      Visibility <- "ST_Maintenance_g_bo_2_Warn_Status_LongDai_HuangYouZui"
      ProcessValue <- "ST_Maintenance_g_u16_2_Times_TiShi_LongDai_HuangYouZui"
   Button "按钮_4" at 606,107 size 196x42; TextOff '1小时后提醒 / 1시간후 다시 알림'
      Visibility <- "ST_Maintenance_g_bo_2_Warn_Status_LongDai_HuangYouZui"
      on Click: ResetBit("ST_Maintenance_g_bo_2_Warn_Status_LongDai_HuangYouZui")
   Button "按钮_5" at 606,156 size 196x42; TextOff '已保养完毕 / 유지보수 이미 완료'; Authorization "User administration"
      Visibility <- "ST_Maintenance_g_bo_2_Warn_Status_LongDai_HuangYouZui"
      on Click: ResetBit("ST_Maintenance_g_bo_2_Status_LongDai_HuangYouZui")
   TextField "文本域_6" at 48,112 size 812x100; Text '保养时间到,请停机第 次为龙带压紧 器加注黄油(耐高温、高速、高负荷) 保养时间到,请停机第 次为龙带压紧 器加注黄油(耐高温、高速、高负荷) 유지보수시간. 기계 스톱. 제 차 tangential belt 압축기에 그리스를 주입한다. (내고온,고속,고부하)'
      Visibility <- "ST_Maintenance_g_bo_3_Warn_Status_LongDai_YaJinQi"
   IOField "IO Field_89" at 355,111 size 70x28; FormatPattern 999
      Visibility <- "ST_Maintenance_g_bo_3_Warn_Status_LongDai_YaJinQi"
      ProcessValue <- "ST_Maintenance_g_u16_3_Times_TiShi_LongDai_YaJinQi"
   Button "按钮_8" at 616,119 size 196x42; TextOff '1小时后提醒 / 1시간후 다시 알림'
      Visibility <- "ST_Maintenance_g_bo_3_Warn_Status_LongDai_YaJinQi"
      on Click: ResetBit("ST_Maintenance_g_bo_3_Warn_Status_LongDai_YaJinQi")
   Button "按钮_9" at 616,168 size 196x42; TextOff '已保养完毕 / 유지보수 이미 완료'; Authorization "User administration"
      Visibility <- "ST_Maintenance_g_bo_3_Warn_Status_LongDai_YaJinQi"
      on Click: ResetBit("ST_Maintenance_g_bo_3_Status_LongDai_YaJinQi")
   TextField "文本域_8" at 32,227 size 812x100; Text '保养时间到,请停机第 次清洗龙带, 注意:水温小于15℃,阴凉通风处晾干,避免日晒 保养时间到,请停机第 次清洗龙带, 注意:水温小于15℃,阴凉通风处晾干,避 免日晒 유지보수시간. 기계 스톱. 제 차 tangential belt를 청소한다. 주의 : 수온이15℃ 이하여야 하며 서늘하고 통풍이 잘 되는곳에 말려야 하며 햇볕에 노출되지 않도 록 해야 한다.'
      Visibility <- "ST_Maintenance_g_bo_5_Warn_Status_LongDai_Clean"
   IOField "IO Field_91" at 338,229 size 70x28; FormatPattern 999
      Visibility <- "ST_Maintenance_g_bo_5_Warn_Status_LongDai_Clean"